(* Logix 5000 project; controller PLC_MCC1201_220AP1 vendor 1 type 14 code 164 rev 35.11; software revision 35.00; part 23 of 25 *)
(* tags used below, declared in another part *)
   xAlwaysOFF : BOOL;
   xAlwaysON : BOOL;
   AUX_xInitialize : BOOL;
   DateTime : DINT[7];   // DINT array tag for retrieve wallclock time through GSV created during conversion
   ForceStatus : INT;   // INT tag to retrieve Force enabled value through GSV created during conversion
   GP_OB_InitializeMain : GP_OB_Initialize;
   GP_OB_InitializeMain_STC : GP_OB_Initialize_STC;
   M2xx_CONVEYOR : MAC_CONVEYOR[20];
   M2xx_CONVEYOR_ALM : MAC_CONVEYOR_ALM[20];
   M2xx_CONVEYOR_HMR : MAC_CONVEYOR_HMR[20];
   M2xx_CONVEYOR_HMW : MAC_CONVEYOR_HMW[20];
   MinorFaultBits : DINT;   // MinorFaultBits
   S : INT[128];
   Status : INT;   // INT tag to retrieve Status value through GSV created during conversion
   TMP_dMacIndex : DINT;
   TMP_xAlwaysOFF : BOOL;
   TMP_xDebugOFF : BOOL;
   Z200 : MAC_Zone_ML;
   Z200_ALM : MAC_Zone_ML_ALM;
   Z200_UPS : ZONE_UPS;
(* MainProgram, continued *)

ROUTINE M2xx_Z200_Conveyors_Faults   (* ladder *)
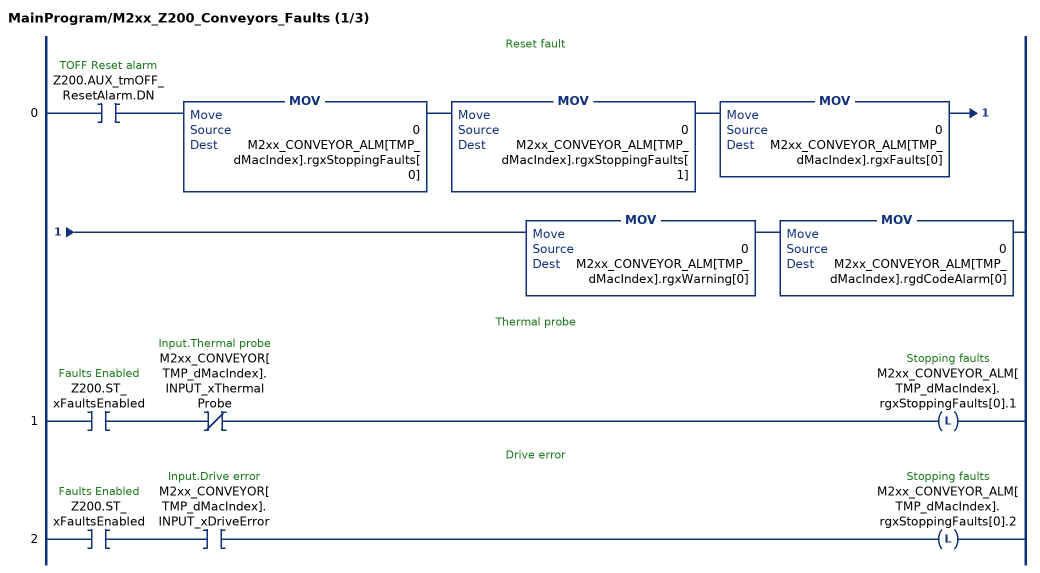
   // Reset fault
   0: XIC(Z200.AUX_tmOFF_ResetAlarm.DN)MOV(0,M2xx_CONVEYOR_ALM[TMP_dMacIndex].rgxStoppingFaults[0])MOV(0,M2xx_CONVEYOR_ALM[TMP_dMacIndex].rgxStoppingFaults[1])MOV(0,M2xx_CONVEYOR_ALM[TMP_dMacIndex].rgxFaults[0])MOV(0,M2xx_CONVEYOR_ALM[TMP_dMacIndex].rgxWarning[0])MOV(0,M2xx_CONVEYOR_ALM[TMP_dMacIndex].rgdCodeAlarm[0]);
   // Thermal probe
   1: XIC(Z200.ST_xFaultsEnabled)XIO(M2xx_CONVEYOR[TMP_dMacIndex].INPUT_xThermalProbe)OTL(M2xx_CONVEYOR_ALM[TMP_dMacIndex].rgxStoppingFaults[0].1);
   // Drive error
   2: XIC(Z200.ST_xFaultsEnabled)XIC(M2xx_CONVEYOR[TMP_dMacIndex].INPUT_xDriveError)OTL(M2xx_CONVEYOR_ALM[TMP_dMacIndex].rgxStoppingFaults[0].2);
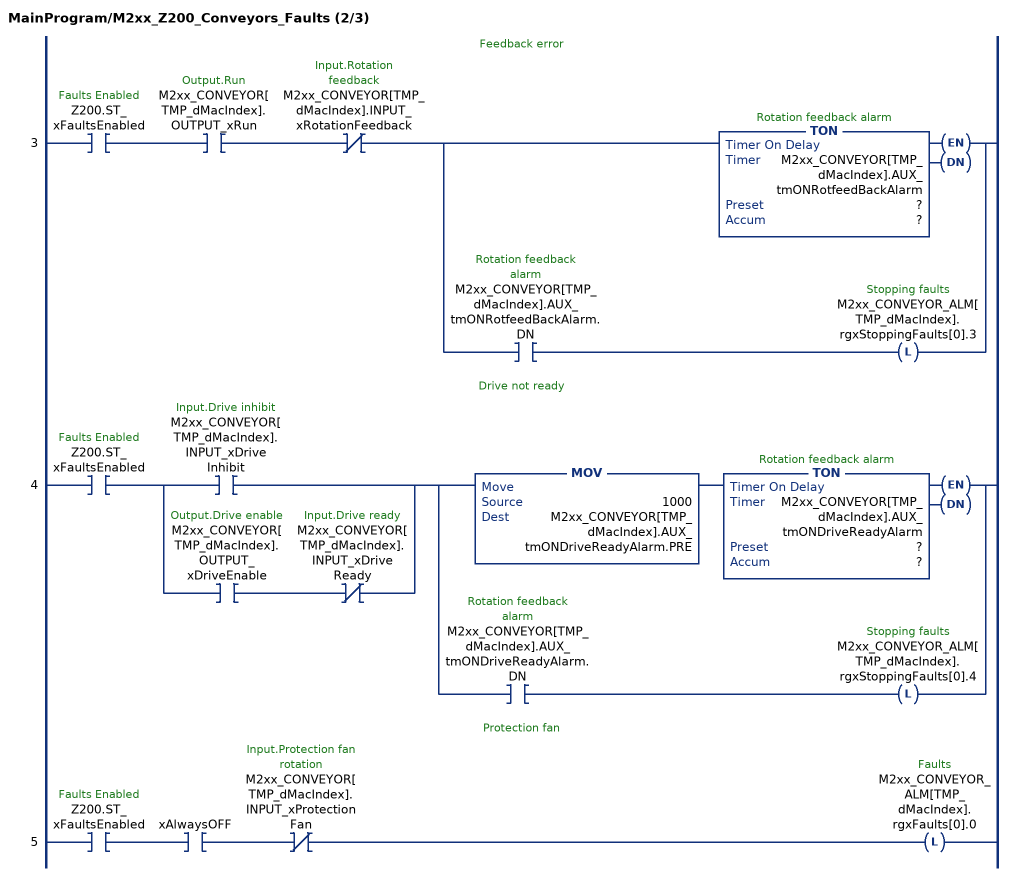
   // Feedback error
   3: XIC(Z200.ST_xFaultsEnabled)XIC(M2xx_CONVEYOR[TMP_dMacIndex].OUTPUT_xRun)XIO(M2xx_CONVEYOR[TMP_dMacIndex].INPUT_xRotationFeedback)[TON(M2xx_CONVEYOR[TMP_dMacIndex].AUX_tmONRotfeedBackAlarm,?,?) ,XIC(M2xx_CONVEYOR[TMP_dMacIndex].AUX_tmONRotfeedBackAlarm.DN) OTL(M2xx_CONVEYOR_ALM[TMP_dMacIndex].rgxStoppingFaults[0].3) ];
   // Drive not ready
   4: XIC(Z200.ST_xFaultsEnabled)[XIC(M2xx_CONVEYOR[TMP_dMacIndex].INPUT_xDriveInhibit) ,XIC(M2xx_CONVEYOR[TMP_dMacIndex].OUTPUT_xDriveEnable) XIO(M2xx_CONVEYOR[TMP_dMacIndex].INPUT_xDriveReady) ][MOV(1000,M2xx_CONVEYOR[TMP_dMacIndex].AUX_tmONDriveReadyAlarm.PRE) TON(M2xx_CONVEYOR[TMP_dMacIndex].AUX_tmONDriveReadyAlarm,?,?) ,XIC(M2xx_CONVEYOR[TMP_dMacIndex].AUX_tmONDriveReadyAlarm.DN) OTL(M2xx_CONVEYOR_ALM[TMP_dMacIndex].rgxStoppingFaults[0].4) ];
   // Protection fan
   5: XIC(Z200.ST_xFaultsEnabled)XIC(xAlwaysOFF)XIO(M2xx_CONVEYOR[TMP_dMacIndex].INPUT_xProtectionFan)OTL(M2xx_CONVEYOR_ALM[TMP_dMacIndex].rgxFaults[0].0);
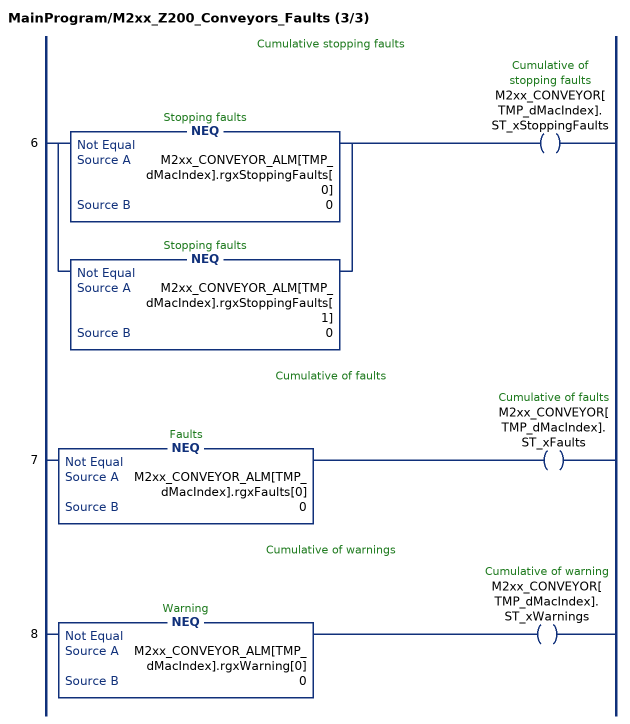
   // Cumulative stopping faults
   6: [NEQ(M2xx_CONVEYOR_ALM[TMP_dMacIndex].rgxStoppingFaults[0],0) ,NEQ(M2xx_CONVEYOR_ALM[TMP_dMacIndex].rgxStoppingFaults[1],0) ]OTE(M2xx_CONVEYOR[TMP_dMacIndex].ST_xStoppingFaults);
   // Cumulative of faults
   7: NEQ(M2xx_CONVEYOR_ALM[TMP_dMacIndex].rgxFaults[0],0)OTE(M2xx_CONVEYOR[TMP_dMacIndex].ST_xFaults);
   // Cumulative of warnings
   8: NEQ(M2xx_CONVEYOR_ALM[TMP_dMacIndex].rgxWarning[0],0)OTE(M2xx_CONVEYOR[TMP_dMacIndex].ST_xWarnings);
END_ROUTINE

ROUTINE M2xx_Z200_Conveyors_Logics   (* ladder *)
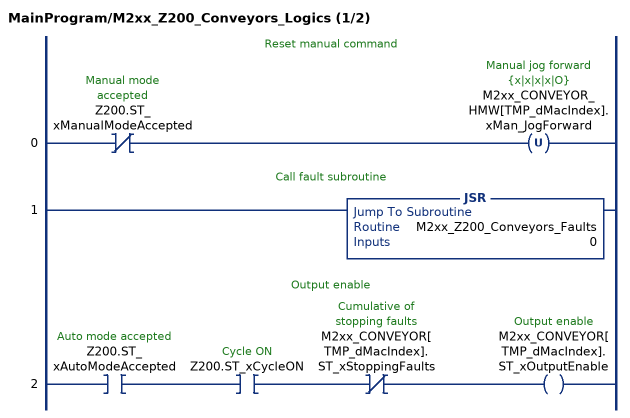
   // Reset manual command
   0: XIO(Z200.ST_xManualModeAccepted)OTU(M2xx_CONVEYOR_HMW[TMP_dMacIndex].xMan_JogForward);
   // Call fault subroutine
   1: JSR(M2xx_Z200_Conveyors_Faults,0);
   // Output enable
   2: XIC(Z200.ST_xAutoModeAccepted)XIC(Z200.ST_xCycleON)XIO(M2xx_CONVEYOR[TMP_dMacIndex].ST_xStoppingFaults)OTE(M2xx_CONVEYOR[TMP_dMacIndex].ST_xOutputEnable);
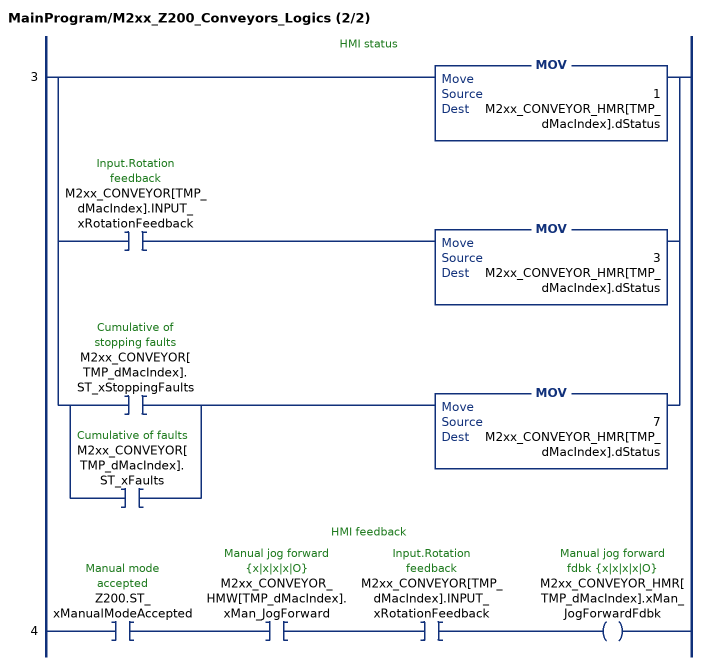
   // HMI status
   3: [MOV(1,M2xx_CONVEYOR_HMR[TMP_dMacIndex].dStatus) ,XIC(M2xx_CONVEYOR[TMP_dMacIndex].INPUT_xRotationFeedback) MOV(3,M2xx_CONVEYOR_HMR[TMP_dMacIndex].dStatus) ,[XIC(M2xx_CONVEYOR[TMP_dMacIndex].ST_xStoppingFaults) ,XIC(M2xx_CONVEYOR[TMP_dMacIndex].ST_xFaults) ] MOV(7,M2xx_CONVEYOR_HMR[TMP_dMacIndex].dStatus) ];
   // HMI feedback
   4: XIC(Z200.ST_xManualModeAccepted)XIC(M2xx_CONVEYOR_HMW[TMP_dMacIndex].xMan_JogForward)XIC(M2xx_CONVEYOR[TMP_dMacIndex].INPUT_xRotationFeedback)OTE(M2xx_CONVEYOR_HMR[TMP_dMacIndex].xMan_JogForwardFdbk);
END_ROUTINE

ROUTINE M2xx_ZUPS_Conveyors_Faults   (* ladder *)
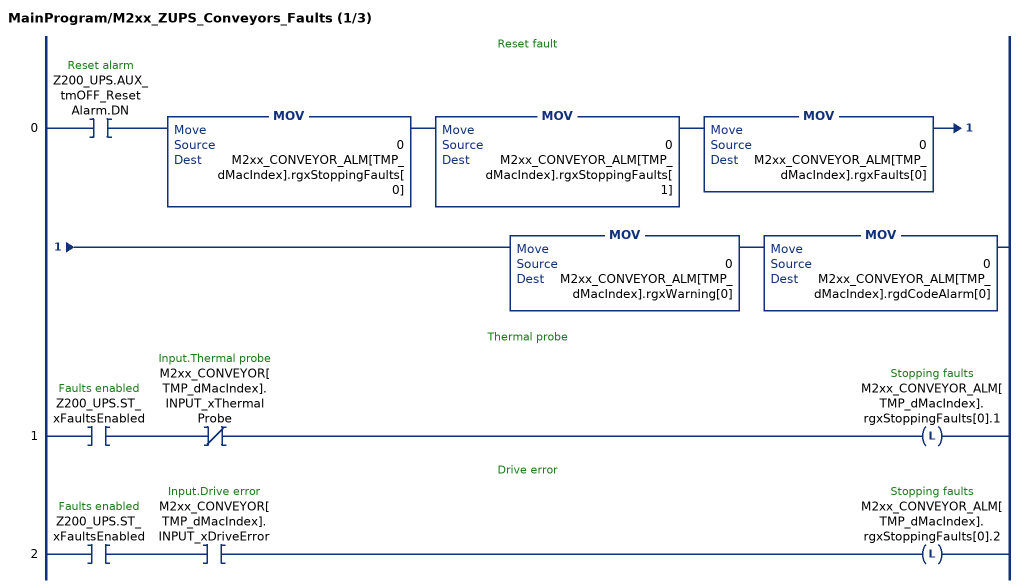
   // Reset fault
   0: XIC(Z200_UPS.AUX_tmOFF_ResetAlarm.DN)MOV(0,M2xx_CONVEYOR_ALM[TMP_dMacIndex].rgxStoppingFaults[0])MOV(0,M2xx_CONVEYOR_ALM[TMP_dMacIndex].rgxStoppingFaults[1])MOV(0,M2xx_CONVEYOR_ALM[TMP_dMacIndex].rgxFaults[0])MOV(0,M2xx_CONVEYOR_ALM[TMP_dMacIndex].rgxWarning[0])MOV(0,M2xx_CONVEYOR_ALM[TMP_dMacIndex].rgdCodeAlarm[0]);
   // Thermal probe
   1: XIC(Z200_UPS.ST_xFaultsEnabled)XIO(M2xx_CONVEYOR[TMP_dMacIndex].INPUT_xThermalProbe)OTL(M2xx_CONVEYOR_ALM[TMP_dMacIndex].rgxStoppingFaults[0].1);
   // Drive error
   2: XIC(Z200_UPS.ST_xFaultsEnabled)XIC(M2xx_CONVEYOR[TMP_dMacIndex].INPUT_xDriveError)OTL(M2xx_CONVEYOR_ALM[TMP_dMacIndex].rgxStoppingFaults[0].2);
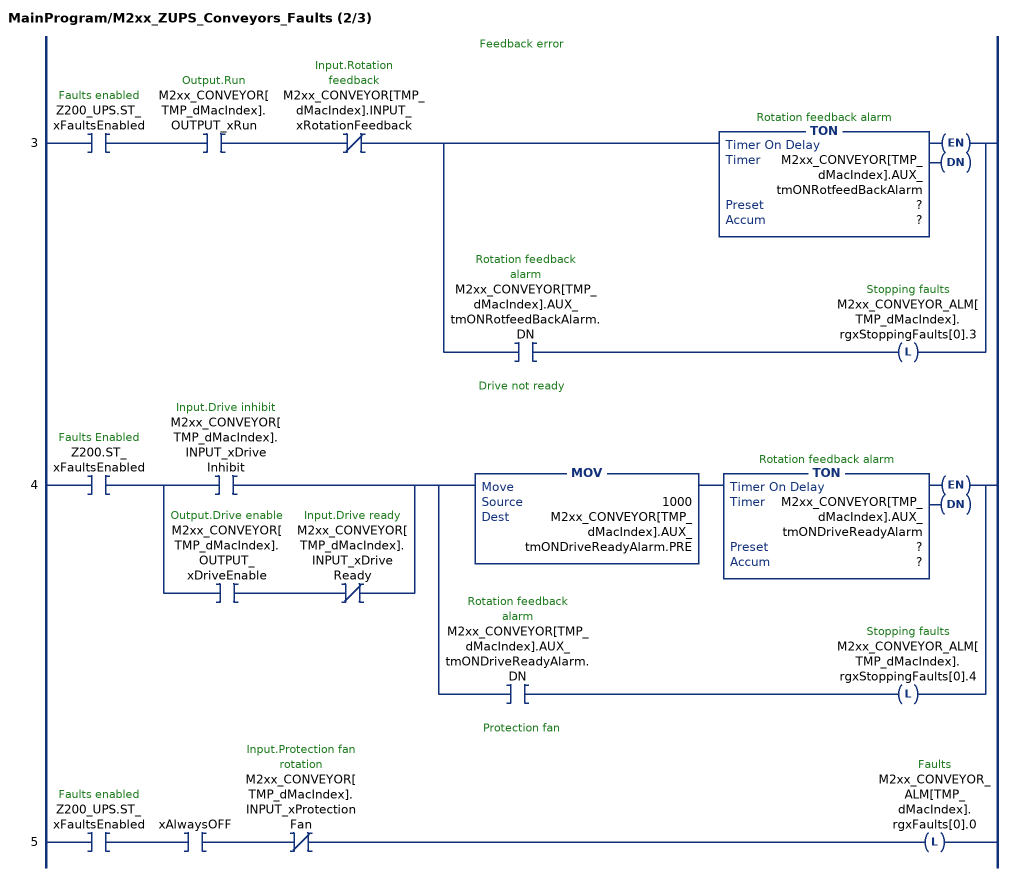
   // Feedback error
   3: XIC(Z200_UPS.ST_xFaultsEnabled)XIC(M2xx_CONVEYOR[TMP_dMacIndex].OUTPUT_xRun)XIO(M2xx_CONVEYOR[TMP_dMacIndex].INPUT_xRotationFeedback)[TON(M2xx_CONVEYOR[TMP_dMacIndex].AUX_tmONRotfeedBackAlarm,?,?) ,XIC(M2xx_CONVEYOR[TMP_dMacIndex].AUX_tmONRotfeedBackAlarm.DN) OTL(M2xx_CONVEYOR_ALM[TMP_dMacIndex].rgxStoppingFaults[0].3) ];
   // Drive not ready
   4: XIC(Z200.ST_xFaultsEnabled)[XIC(M2xx_CONVEYOR[TMP_dMacIndex].INPUT_xDriveInhibit) ,XIC(M2xx_CONVEYOR[TMP_dMacIndex].OUTPUT_xDriveEnable) XIO(M2xx_CONVEYOR[TMP_dMacIndex].INPUT_xDriveReady) ][MOV(1000,M2xx_CONVEYOR[TMP_dMacIndex].AUX_tmONDriveReadyAlarm.PRE) TON(M2xx_CONVEYOR[TMP_dMacIndex].AUX_tmONDriveReadyAlarm,?,?) ,XIC(M2xx_CONVEYOR[TMP_dMacIndex].AUX_tmONDriveReadyAlarm.DN) OTL(M2xx_CONVEYOR_ALM[TMP_dMacIndex].rgxStoppingFaults[0].4) ];
   // Protection fan
   5: XIC(Z200_UPS.ST_xFaultsEnabled)XIC(xAlwaysOFF)XIO(M2xx_CONVEYOR[TMP_dMacIndex].INPUT_xProtectionFan)OTL(M2xx_CONVEYOR_ALM[TMP_dMacIndex].rgxFaults[0].0);
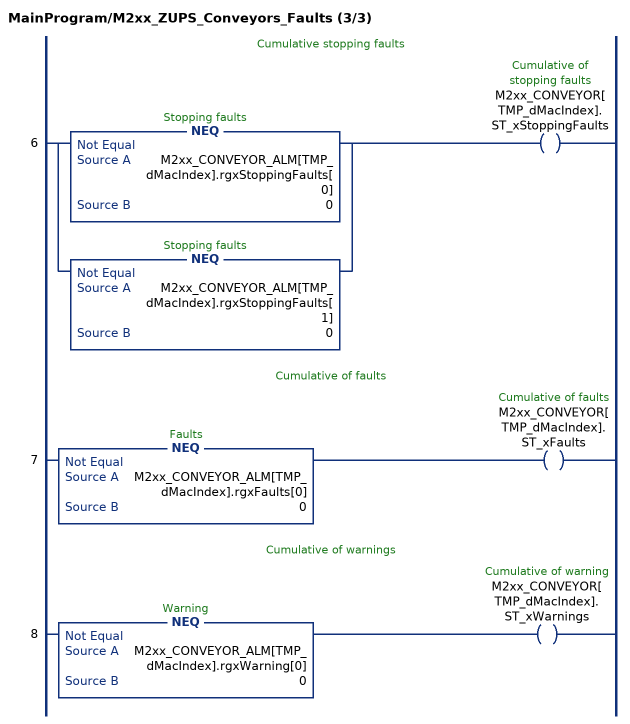
   // Cumulative stopping faults
   6: [NEQ(M2xx_CONVEYOR_ALM[TMP_dMacIndex].rgxStoppingFaults[0],0) ,NEQ(M2xx_CONVEYOR_ALM[TMP_dMacIndex].rgxStoppingFaults[1],0) ]OTE(M2xx_CONVEYOR[TMP_dMacIndex].ST_xStoppingFaults);
   // Cumulative of faults
   7: NEQ(M2xx_CONVEYOR_ALM[TMP_dMacIndex].rgxFaults[0],0)OTE(M2xx_CONVEYOR[TMP_dMacIndex].ST_xFaults);
   // Cumulative of warnings
   8: NEQ(M2xx_CONVEYOR_ALM[TMP_dMacIndex].rgxWarning[0],0)OTE(M2xx_CONVEYOR[TMP_dMacIndex].ST_xWarnings);
END_ROUTINE

ROUTINE M2xx_ZUPS_Conveyors_Logics   (* ladder *)
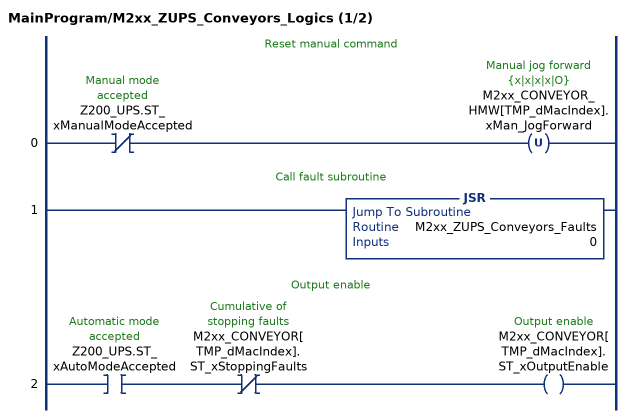
   // Reset manual command
   0: XIO(Z200_UPS.ST_xManualModeAccepted)OTU(M2xx_CONVEYOR_HMW[TMP_dMacIndex].xMan_JogForward);
   // Call fault subroutine
   1: JSR(M2xx_ZUPS_Conveyors_Faults,0);
   // Output enable
   2: XIC(Z200_UPS.ST_xAutoModeAccepted)XIO(M2xx_CONVEYOR[TMP_dMacIndex].ST_xStoppingFaults)OTE(M2xx_CONVEYOR[TMP_dMacIndex].ST_xOutputEnable);
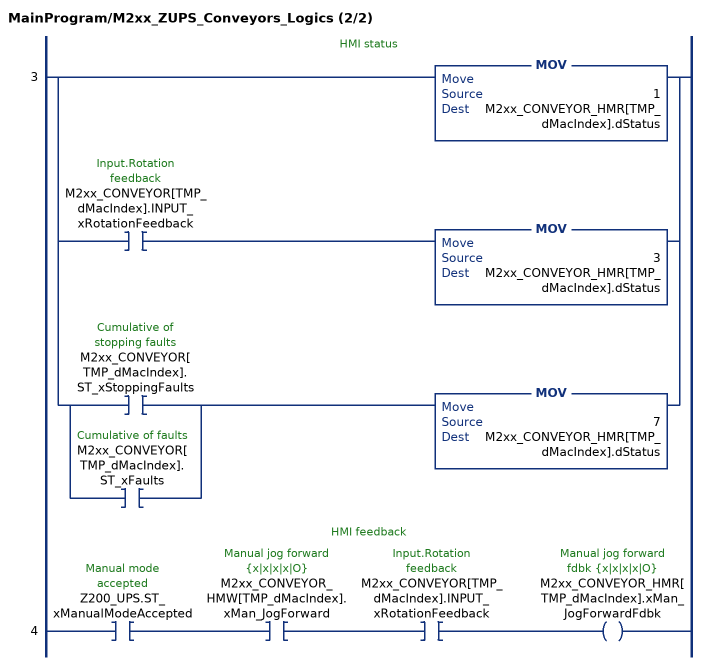
   // HMI status
   3: [MOV(1,M2xx_CONVEYOR_HMR[TMP_dMacIndex].dStatus) ,XIC(M2xx_CONVEYOR[TMP_dMacIndex].INPUT_xRotationFeedback) MOV(3,M2xx_CONVEYOR_HMR[TMP_dMacIndex].dStatus) ,[XIC(M2xx_CONVEYOR[TMP_dMacIndex].ST_xStoppingFaults) ,XIC(M2xx_CONVEYOR[TMP_dMacIndex].ST_xFaults) ] MOV(7,M2xx_CONVEYOR_HMR[TMP_dMacIndex].dStatus) ];
   // HMI feedback
   4: XIC(Z200_UPS.ST_xManualModeAccepted)XIC(M2xx_CONVEYOR_HMW[TMP_dMacIndex].xMan_JogForward)XIC(M2xx_CONVEYOR[TMP_dMacIndex].INPUT_xRotationFeedback)OTE(M2xx_CONVEYOR_HMR[TMP_dMacIndex].xMan_JogForwardFdbk);
END_ROUTINE

ROUTINE MainRoutine   (* ladder *)
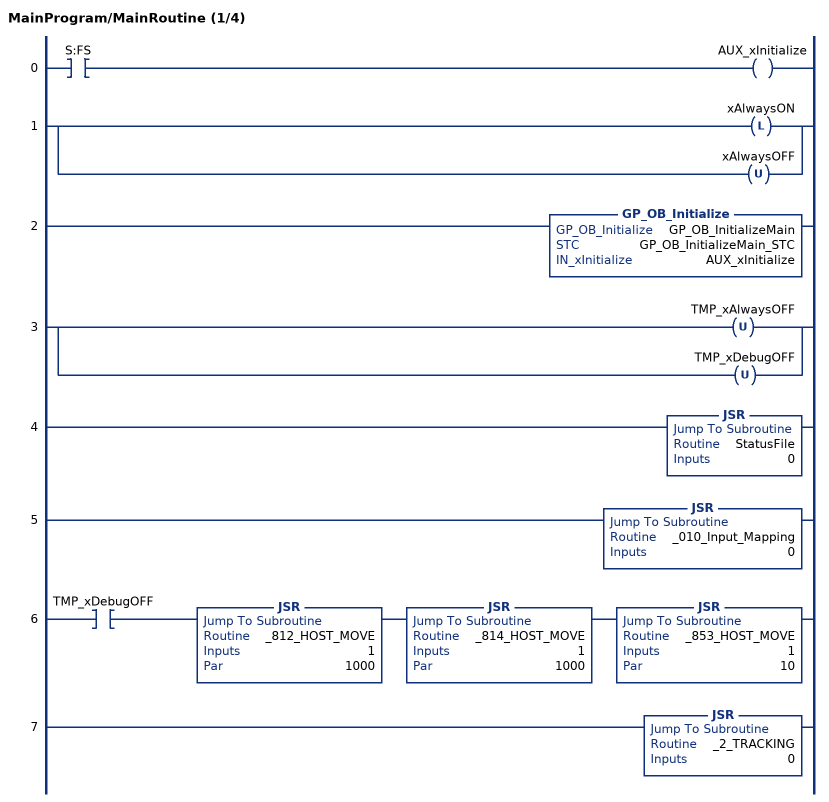
   0: XIC(S:FS)OTE(AUX_xInitialize);
   1: [OTL(xAlwaysON) ,OTU(xAlwaysOFF) ];
   2: GP_OB_Initialize(GP_OB_InitializeMain,GP_OB_InitializeMain_STC,AUX_xInitialize);
   3: [OTU(TMP_xAlwaysOFF) ,OTU(TMP_xDebugOFF) ];
   4: JSR(StatusFile,0);
   5: JSR(_010_Input_Mapping,0);
   6: XIC(TMP_xDebugOFF)JSR(_812_HOST_MOVE,1,1000)JSR(_814_HOST_MOVE,1,1000)JSR(_853_HOST_MOVE,1,10);
   7: JSR(_2_TRACKING,0);
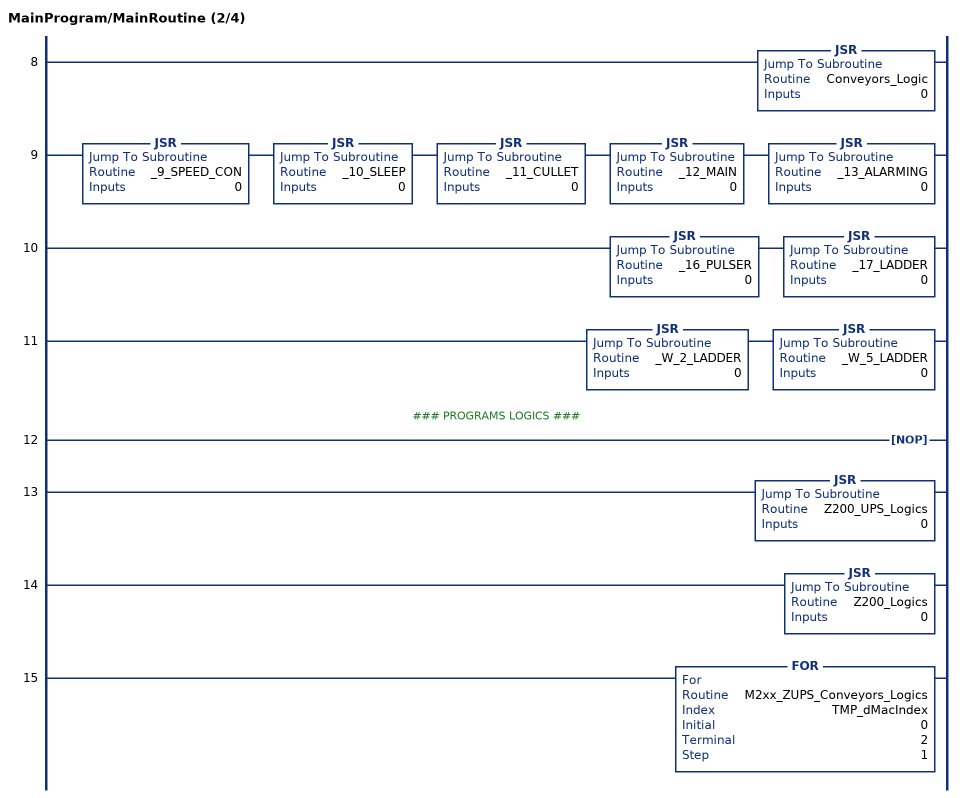
   8: JSR(Conveyors_Logic,0);
   9: JSR(_9_SPEED_CON,0)JSR(_10_SLEEP,0)JSR(_11_CULLET,0)JSR(_12_MAIN,0)JSR(_13_ALARMING,0);
   10: JSR(_16_PULSER,0)JSR(_17_LADDER,0);
   11: JSR(_W_2_LADDER,0)JSR(_W_5_LADDER,0);
   // ### PROGRAMS LOGICS ###
   12: NOP();
   13: JSR(Z200_UPS_Logics,0);
   14: JSR(Z200_Logics,0);
   15: FOR(M2xx_ZUPS_Conveyors_Logics,TMP_dMacIndex,0,2,1);
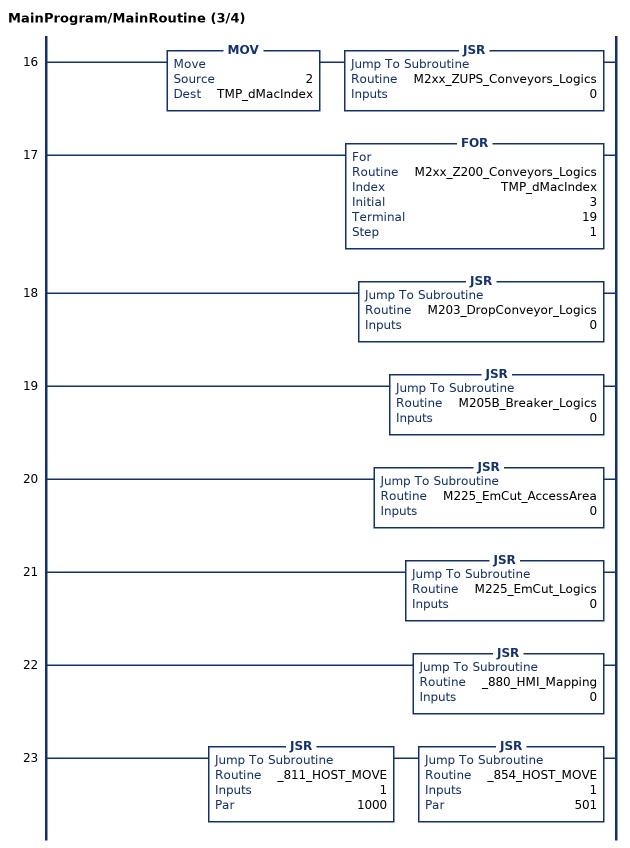
   16: MOV(2,TMP_dMacIndex)JSR(M2xx_ZUPS_Conveyors_Logics,0);
   17: FOR(M2xx_Z200_Conveyors_Logics,TMP_dMacIndex,3,19,1);
   18: JSR(M203_DropConveyor_Logics,0);
   19: JSR(M205B_Breaker_Logics,0);
   20: JSR(M225_EmCut_AccessArea,0);
   21: JSR(M225_EmCut_Logics,0);
   22: JSR(_880_HMI_Mapping,0);
   23: JSR(_811_HOST_MOVE,1,1000)JSR(_854_HOST_MOVE,1,501);
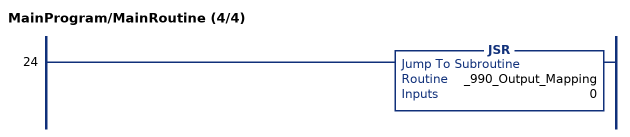
   24: JSR(_990_Output_Mapping,0);
END_ROUTINE

ROUTINE StatusFile   (* ladder *)
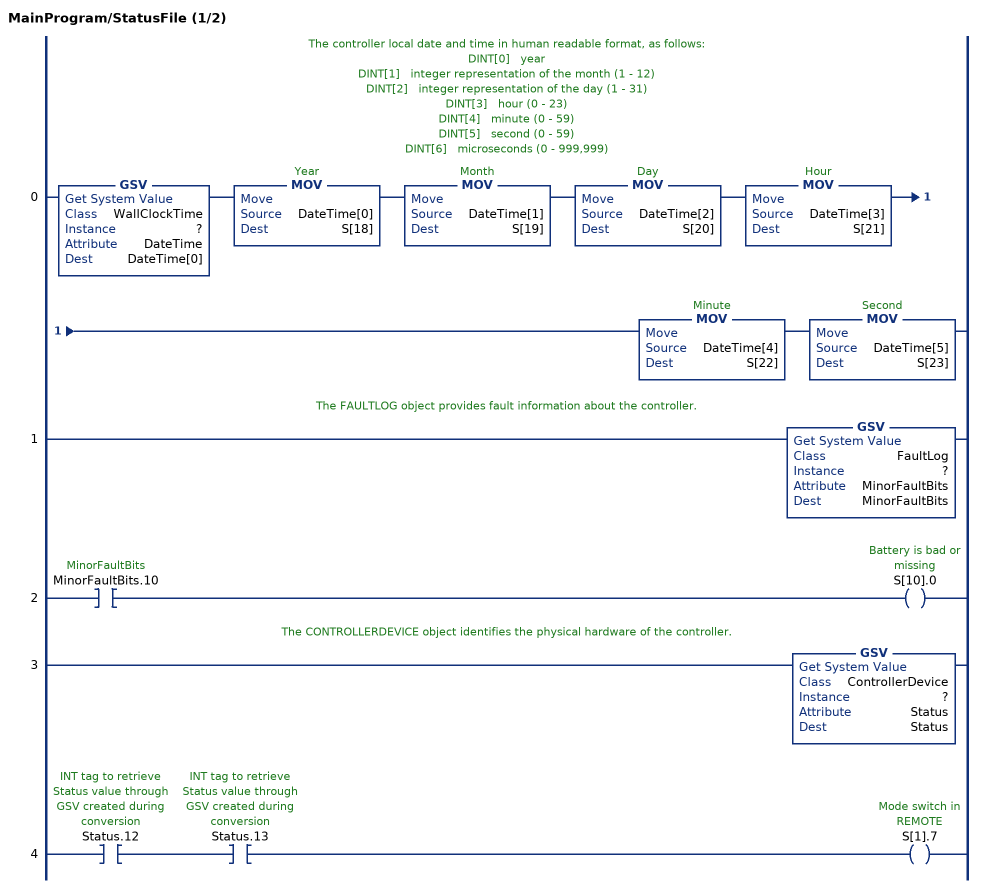
   // The controller local date and time in human readable format, as follows:
   // DINT[0] 	year
   // DINT[1] 	integer representation of the month (1 - 12)
   // DINT[2] 	integer representation of the day (1 - 31)
   // DINT[3] 	hour (0 - 23)
   // DINT[4] 	minute (0 - 59)
   // DINT[5] 	second (0 - 59)
   // DINT[6] 	microseconds (0 - 999,999)
   0: GSV(WallClockTime,?,DateTime,DateTime[0])MOV(DateTime[0],S[18])MOV(DateTime[1],S[19])MOV(DateTime[2],S[20])MOV(DateTime[3],S[21])MOV(DateTime[4],S[22])MOV(DateTime[5],S[23]);
   // The FAULTLOG object provides fault information about the controller.
   1: GSV(FaultLog,?,MinorFaultBits,MinorFaultBits);
   2: XIC(MinorFaultBits.10)OTE(S[10].0);
   // The CONTROLLERDEVICE object identifies the physical hardware of the controller.
   3: GSV(ControllerDevice,?,Status,Status);
   4: XIC(Status.12)XIC(Status.13)OTE(S[1].7);
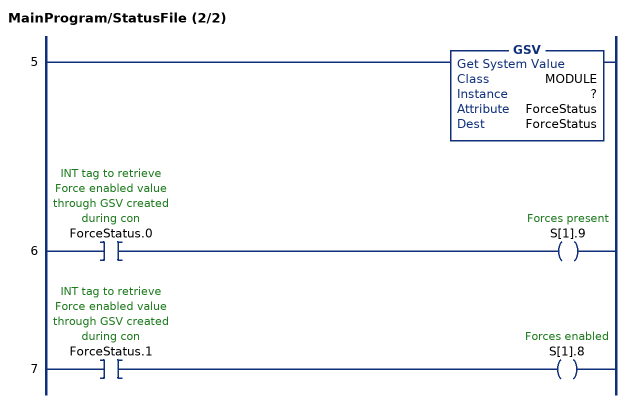
   5: GSV(MODULE,?,ForceStatus,ForceStatus);
   6: XIC(ForceStatus.0)OTE(S[1].9);
   7: XIC(ForceStatus.1)OTE(S[1].8);
END_ROUTINE

ROUTINE Z200_Faults   (* ladder *)
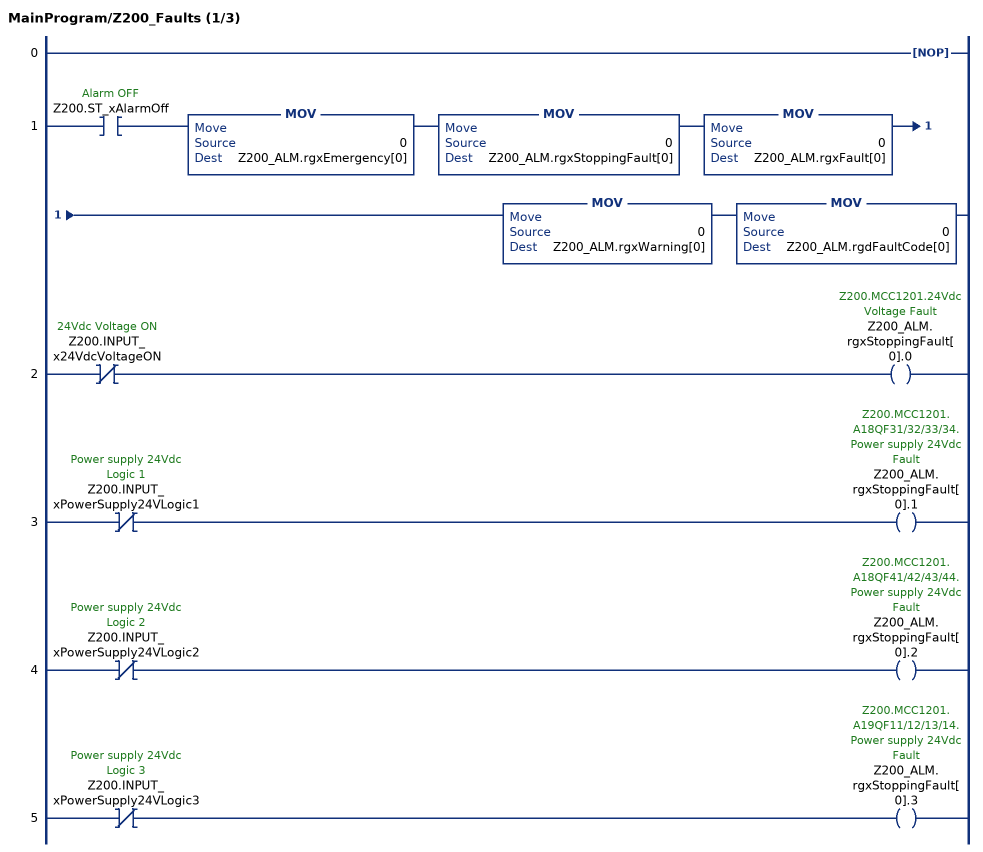
   0: NOP();
   1: XIC(Z200.ST_xAlarmOff)MOV(0,Z200_ALM.rgxEmergency[0])MOV(0,Z200_ALM.rgxStoppingFault[0])MOV(0,Z200_ALM.rgxFault[0])MOV(0,Z200_ALM.rgxWarning[0])MOV(0,Z200_ALM.rgdFaultCode[0]);
   2: XIO(Z200.INPUT_x24VdcVoltageON)OTE(Z200_ALM.rgxStoppingFault[0].0);
   3: XIO(Z200.INPUT_xPowerSupply24VLogic1)OTE(Z200_ALM.rgxStoppingFault[0].1);
   4: XIO(Z200.INPUT_xPowerSupply24VLogic2)OTE(Z200_ALM.rgxStoppingFault[0].2);
   5: XIO(Z200.INPUT_xPowerSupply24VLogic3)OTE(Z200_ALM.rgxStoppingFault[0].3);
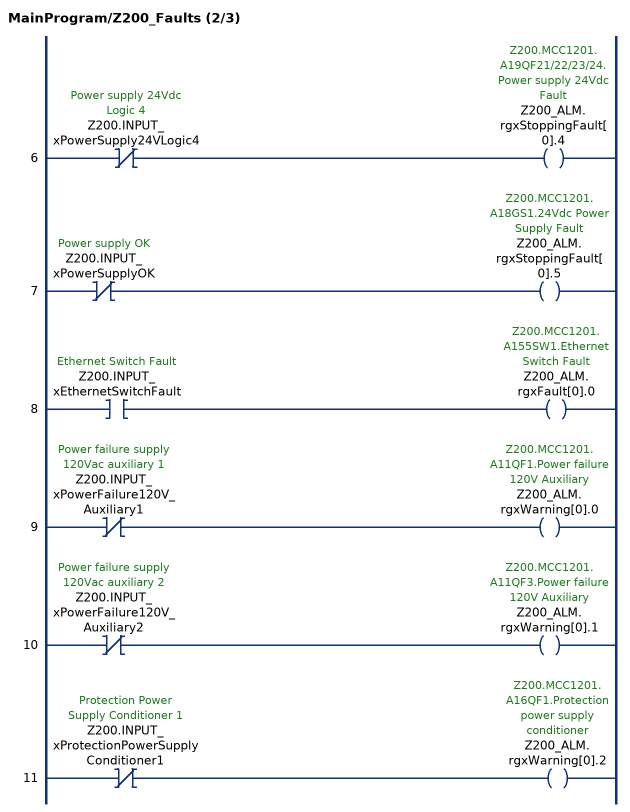
   6: XIO(Z200.INPUT_xPowerSupply24VLogic4)OTE(Z200_ALM.rgxStoppingFault[0].4);
   7: XIO(Z200.INPUT_xPowerSupplyOK)OTE(Z200_ALM.rgxStoppingFault[0].5);
   8: XIC(Z200.INPUT_xEthernetSwitchFault)OTE(Z200_ALM.rgxFault[0].0);
   9: XIO(Z200.INPUT_xPowerFailure120V_Auxiliary1)OTE(Z200_ALM.rgxWarning[0].0);
   10: XIO(Z200.INPUT_xPowerFailure120V_Auxiliary2)OTE(Z200_ALM.rgxWarning[0].1);
   11: XIO(Z200.INPUT_xProtectionPowerSupplyConditioner1)OTE(Z200_ALM.rgxWarning[0].2);
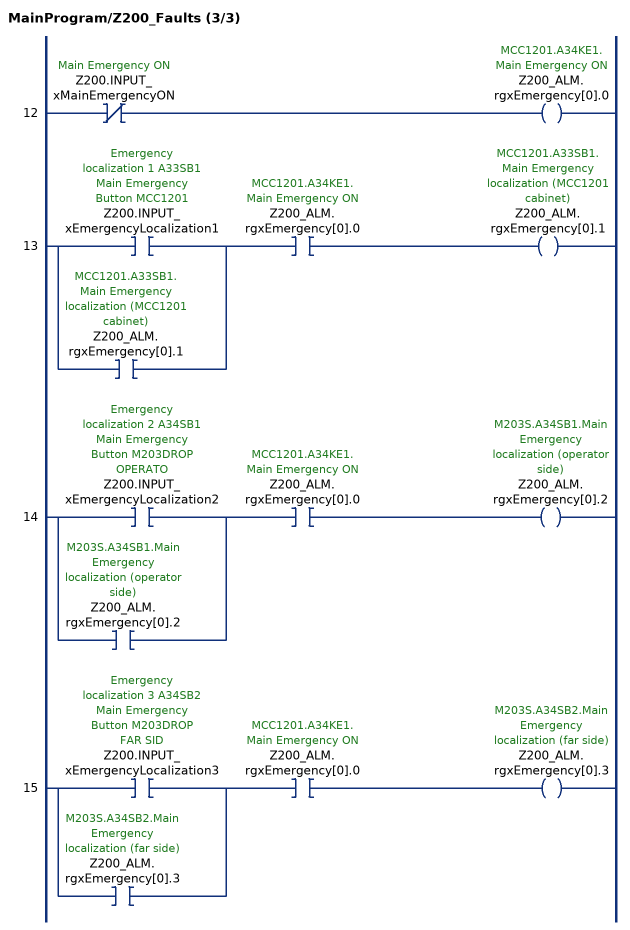
   12: XIO(Z200.INPUT_xMainEmergencyON)OTE(Z200_ALM.rgxEmergency[0].0);
   13: [XIC(Z200.INPUT_xEmergencyLocalization1) ,XIC(Z200_ALM.rgxEmergency[0].1) ]XIC(Z200_ALM.rgxEmergency[0].0)OTE(Z200_ALM.rgxEmergency[0].1);
   14: [XIC(Z200.INPUT_xEmergencyLocalization2) ,XIC(Z200_ALM.rgxEmergency[0].2) ]XIC(Z200_ALM.rgxEmergency[0].0)OTE(Z200_ALM.rgxEmergency[0].2);
   15: [XIC(Z200.INPUT_xEmergencyLocalization3) ,XIC(Z200_ALM.rgxEmergency[0].3) ]XIC(Z200_ALM.rgxEmergency[0].0)OTE(Z200_ALM.rgxEmergency[0].3);
END_ROUTINE
